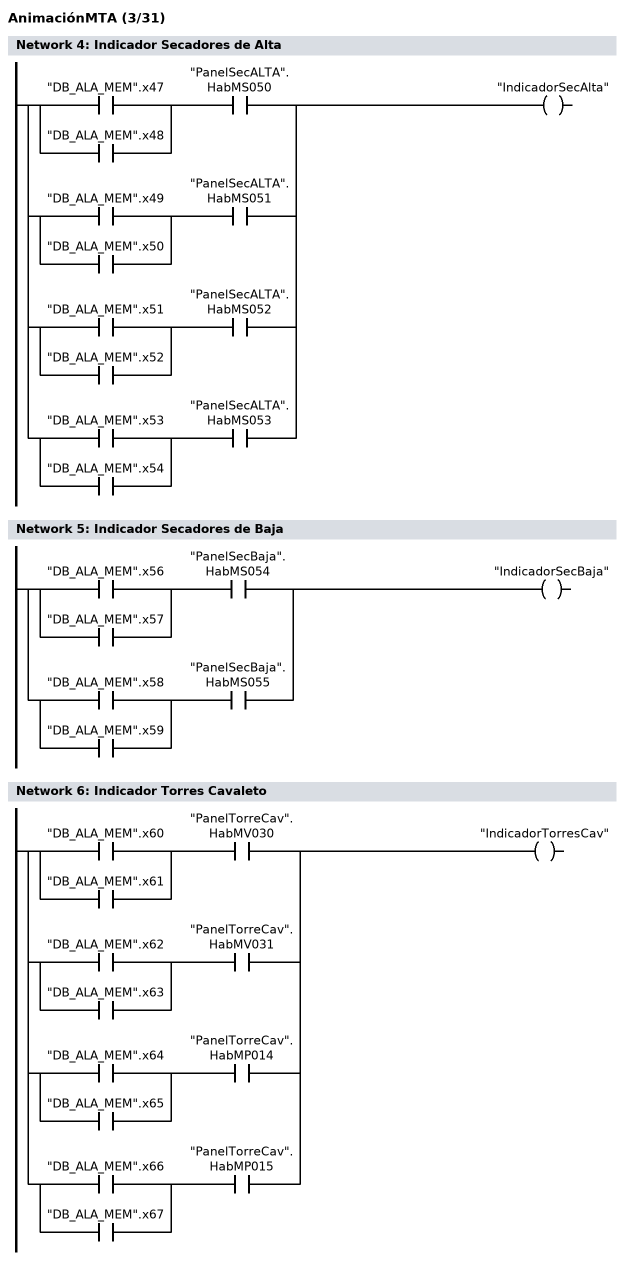
   RUNG wire#powerrail
      Contact( "DB_ALA_MEM".x47 )
      wire#w1
      Contact( "PanelSecALTA".HabMS050 )
      wire#w2
      Coil( "IndicadorSecAlta" )
   END_RUNG
   RUNG wire#powerrail
      Contact( "DB_ALA_MEM".x48 )
   END_RUNG wire#w1
   RUNG wire#powerrail
      Contact( "DB_ALA_MEM".x49 )
      wire#w3
      Contact( "PanelSecALTA".HabMS051 )
   END_RUNG wire#w2
   RUNG wire#powerrail
      Contact( "DB_ALA_MEM".x50 )
   END_RUNG wire#w3
   RUNG wire#powerrail
      Contact( "DB_ALA_MEM".x51 )
      wire#w4
      Contact( "PanelSecALTA".HabMS052 )
   END_RUNG wire#w2
   RUNG wire#powerrail
      Contact( "DB_ALA_MEM".x52 )
   END_RUNG wire#w4
   RUNG wire#powerrail
      Contact( "DB_ALA_MEM".x53 )
      wire#w5
      Contact( "PanelSecALTA".HabMS053 )
   END_RUNG wire#w2
   RUNG wire#powerrail
      Contact( "DB_ALA_MEM".x54 )
   END_RUNG wire#w5
   // the same network as SCL:
   "IndicadorSecAlta" := (("DB_ALA_MEM".x47 OR "DB_ALA_MEM".x48) AND "PanelSecALTA".HabMS050) OR (("DB_ALA_MEM".x49 OR "DB_ALA_MEM".x50) AND "PanelSecALTA".HabMS051) OR (("DB_ALA_MEM".x51 OR "DB_ALA_MEM".x52) AND "PanelSecALTA".HabMS052) OR (("DB_ALA_MEM".x53 OR "DB_ALA_MEM".x54) AND "PanelSecALTA".HabMS053);
END_REGION

REGION Network 5: Indicador Secadores de Baja
   RUNG wire#powerrail
      Contact( "DB_ALA_MEM".x56 )
      wire#w1
      Contact( "PanelSecBaja".HabMS054 )
      wire#w2
      Coil( "IndicadorSecBaja" )
   END_RUNG
   RUNG wire#powerrail
      Contact( "DB_ALA_MEM".x57 )
   END_RUNG wire#w1
   RUNG wire#powerrail
      Contact( "DB_ALA_MEM".x58 )
      wire#w3
      Contact( "PanelSecBaja".HabMS055 )
   END_RUNG wire#w2
   RUNG wire#powerrail
      Contact( "DB_ALA_MEM".x59 )
   END_RUNG wire#w3
   // the same network as SCL:
   "IndicadorSecBaja" := (("DB_ALA_MEM".x56 OR "DB_ALA_MEM".x57) AND "PanelSecBaja".HabMS054) OR (("DB_ALA_MEM".x58 OR "DB_ALA_MEM".x59) AND "PanelSecBaja".HabMS055);
END_REGION

REGION Network 6: Indicador Torres Cavaleto
   RUNG wire#powerrail
      Contact( "DB_ALA_MEM".x60 )
      wire#w1
      Contact( "PanelTorreCav".HabMV030 )
      wire#w2
      Coil( "IndicadorTorresCav" )
   END_RUNG
   RUNG wire#powerrail
      Contact( "DB_ALA_MEM".x61 )
   END_RUNG wire#w1
   RUNG wire#powerrail
      Contact( "DB_ALA_MEM".x62 )
      wire#w3
      Contact( "PanelTorreCav".HabMV031 )
   END_RUNG wire#w2
   RUNG wire#powerrail
      Contact( "DB_ALA_MEM".x63 )
   END_RUNG wire#w3
   RUNG wire#powerrail
      Contact( "DB_ALA_MEM".x64 )
      wire#w4
      Contact( "PanelTorreCav".HabMP014 )
   END_RUNG wire#w2
   RUNG wire#powerrail
      Contact( "DB_ALA_MEM".x65 )
   END_RUNG wire#w4
   RUNG wire#powerrail
      Contact( "DB_ALA_MEM".x66 )
      wire#w5
      Contact( "PanelTorreCav".HabMP015 )
   END_RUNG wire#w2
   RUNG wire#powerrail
      Contact( "DB_ALA_MEM".x67 )
   END_RUNG wire#w5
   // the same network as SCL:
   "IndicadorTorresCav" := (("DB_ALA_MEM".x60 OR "DB_ALA_MEM".x61) AND "PanelTorreCav".HabMV030) OR (("DB_ALA_MEM".x62 OR "DB_ALA_MEM".x63) AND "PanelTorreCav".HabMV031) OR (("DB_ALA_MEM".x64 OR "DB_ALA_MEM".x65) AND "PanelTorreCav".HabMP014) OR (("DB_ALA_MEM".x66 OR "DB_ALA_MEM".x67) AND "PanelTorreCav".HabMP015);
END_REGION

REGION Network 7: Indicador Compresores de Alta
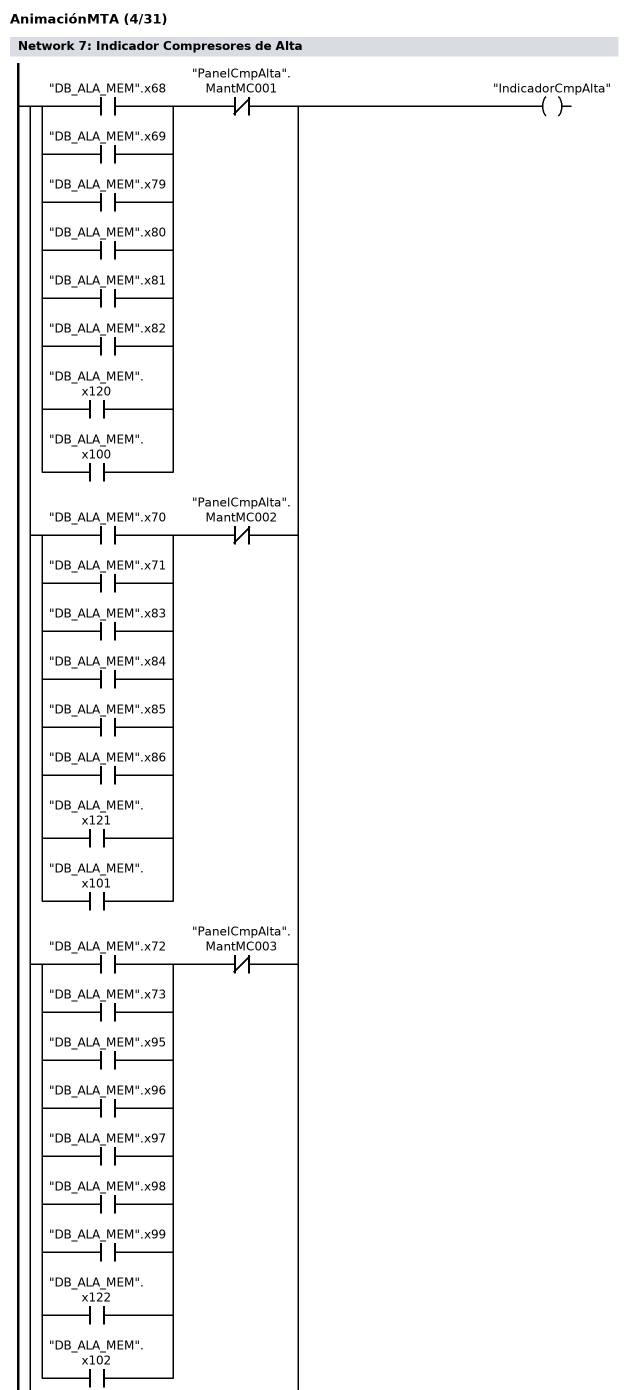
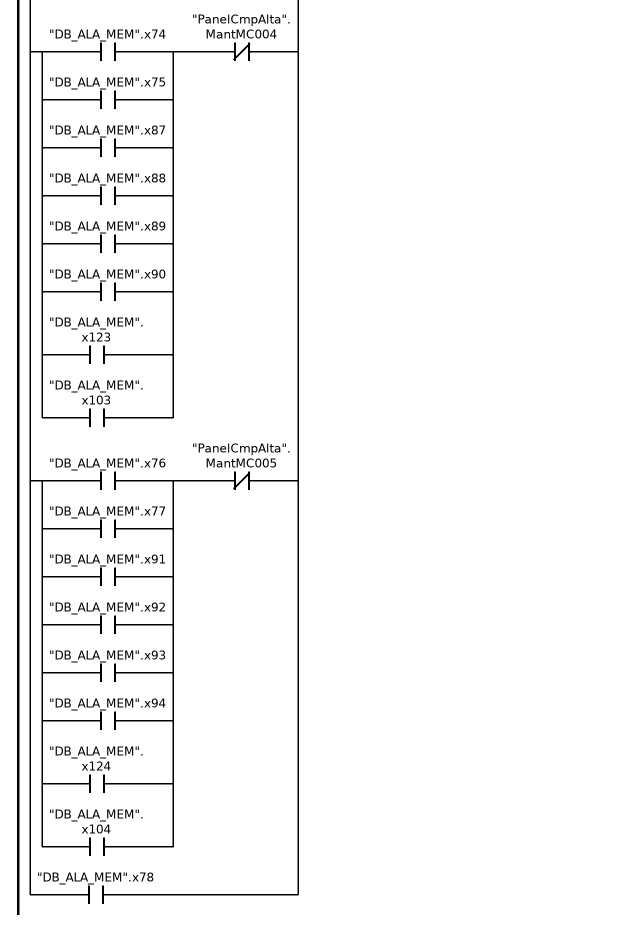
   RUNG wire#powerrail
      Contact( "DB_ALA_MEM".x68 )
      wire#w1
      I_Contact( "PanelCmpAlta".MantMC001 )
      wire#w2
      Coil( "IndicadorCmpAlta" )
   END_RUNG
   RUNG wire#powerrail
      Contact( "DB_ALA_MEM".x69 )
   END_RUNG wire#w1
   RUNG wire#powerrail
      Contact( "DB_ALA_MEM".x79 )
   END_RUNG wire#w1
   RUNG wire#powerrail
      Contact( "DB_ALA_MEM".x80 )
   END_RUNG wire#w1
   RUNG wire#powerrail
      Contact( "DB_ALA_MEM".x81 )
   END_RUNG wire#w1
   RUNG wire#powerrail
      Contact( "DB_ALA_MEM".x82 )
   END_RUNG wire#w1
   RUNG wire#powerrail
      Contact( "DB_ALA_MEM".x120 )
   END_RUNG wire#w1
   RUNG wire#powerrail
      Contact( "DB_ALA_MEM".x100 )
   END_RUNG wire#w1
   RUNG wire#powerrail
      Contact( "DB_ALA_MEM".x70 )
      wire#w3
      I_Contact( "PanelCmpAlta".MantMC002 )
   END_RUNG wire#w2
   RUNG wire#powerrail
      Contact( "DB_ALA_MEM".x71 )
   END_RUNG wire#w3
   RUNG wire#powerrail
      Contact( "DB_ALA_MEM".x83 )
   END_RUNG wire#w3
   RUNG wire#powerrail
      Contact( "DB_ALA_MEM".x84 )
   END_RUNG wire#w3
   RUNG wire#powerrail
      Contact( "DB_ALA_MEM".x85 )
   END_RUNG wire#w3
   RUNG wire#powerrail
      Contact( "DB_ALA_MEM".x86 )
   END_RUNG wire#w3
   RUNG wire#powerrail
      Contact( "DB_ALA_MEM".x121 )
   END_RUNG wire#w3
   RUNG wire#powerrail
      Contact( "DB_ALA_MEM".x101 )
   END_RUNG wire#w3
   RUNG wire#powerrail
      Contact( "DB_ALA_MEM".x72 )
      wire#w4
      I_Contact( "PanelCmpAlta".MantMC003 )
   END_RUNG wire#w2
   RUNG wire#powerrail
      Contact( "DB_ALA_MEM".x73 )
   END_RUNG wire#w4
   RUNG wire#powerrail
      Contact( "DB_ALA_MEM".x95 )
   END_RUNG wire#w4
   RUNG wire#powerrail
      Contact( "DB_ALA_MEM".x96 )
   END_RUNG wire#w4
   RUNG wire#powerrail
      Contact( "DB_ALA_MEM".x97 )
   END_RUNG wire#w4
   RUNG wire#powerrail
      Contact( "DB_ALA_MEM".x98 )
   END_RUNG wire#w4
   RUNG wire#powerrail
      Contact( "DB_ALA_MEM".x99 )
   END_RUNG wire#w4
   RUNG wire#powerrail
      Contact( "DB_ALA_MEM".x122 )
   END_RUNG wire#w4
   RUNG wire#powerrail
      Contact( "DB_ALA_MEM".x102 )
   END_RUNG wire#w4
   RUNG wire#powerrail
      Contact( "DB_ALA_MEM".x74 )
      wire#w5
      I_Contact( "PanelCmpAlta".MantMC004 )
   END_RUNG wire#w2
   RUNG wire#powerrail
      Contact( "DB_ALA_MEM".x75 )
   END_RUNG wire#w5
   RUNG wire#powerrail
      Contact( "DB_ALA_MEM".x87 )
   END_RUNG wire#w5
   RUNG wire#powerrail
      Contact( "DB_ALA_MEM".x88 )
   END_RUNG wire#w5
   RUNG wire#powerrail
      Contact( "DB_ALA_MEM".x89 )
   END_RUNG wire#w5
   RUNG wire#powerrail
      Contact( "DB_ALA_MEM".x90 )
   END_RUNG wire#w5
   RUNG wire#powerrail
      Contact( "DB_ALA_MEM".x123 )
   END_RUNG wire#w5
   RUNG wire#powerrail
      Contact( "DB_ALA_MEM".x103 )
   END_RUNG wire#w5
   RUNG wire#powerrail
      Contact( "DB_ALA_MEM".x76 )
      wire#w6
      I_Contact( "PanelCmpAlta".MantMC005 )
   END_RUNG wire#w2
   RUNG wire#powerrail
      Contact( "DB_ALA_MEM".x77 )
   END_RUNG wire#w6
   RUNG wire#powerrail
      Contact( "DB_ALA_MEM".x91 )
   END_RUNG wire#w6
   RUNG wire#powerrail
      Contact( "DB_ALA_MEM".x92 )
   END_RUNG wire#w6
   RUNG wire#powerrail
      Contact( "DB_ALA_MEM".x93 )
   END_RUNG wire#w6
   RUNG wire#powerrail
      Contact( "DB_ALA_MEM".x94 )
   END_RUNG wire#w6
   RUNG wire#powerrail
      Contact( "DB_ALA_MEM".x124 )
   END_RUNG wire#w6
   RUNG wire#powerrail
      Contact( "DB_ALA_MEM".x104 )
   END_RUNG wire#w6
   RUNG wire#powerrail
      Contact( "DB_ALA_MEM".x78 )
   END_RUNG wire#w2
   // the same network as SCL:
   "IndicadorCmpAlta" := (("DB_ALA_MEM".x68 OR "DB_ALA_MEM".x69 OR "DB_ALA_MEM".x79 OR "DB_ALA_MEM".x80 OR "DB_ALA_MEM".x81 OR "DB_ALA_MEM".x82 OR "DB_ALA_MEM".x120 OR "DB_ALA_MEM".x100) AND NOT "PanelCmpAlta".MantMC001) OR (("DB_ALA_MEM".x70 OR "DB_ALA_MEM".x71 OR "DB_ALA_MEM".x83 OR "DB_ALA_MEM".x84 OR "DB_ALA_MEM".x85 OR "DB_ALA_MEM".x86 OR "DB_ALA_MEM".x121 OR "DB_ALA_MEM".x101) AND NOT "PanelCmpAlta".MantMC002) OR (("DB_ALA_MEM".x72 OR "DB_ALA_MEM".x73 OR "DB_ALA_MEM".x95 OR "DB_ALA_MEM".x96 OR "DB_ALA_MEM".x97 OR "DB_ALA_MEM".x98 OR "DB_ALA_MEM".x99 OR "DB_ALA_MEM".x122 OR "DB_ALA_MEM".x102) AND NOT "PanelCmpAlta".MantMC003) OR (("DB_ALA_MEM".x74 OR "DB_ALA_MEM".x75 OR "DB_ALA_MEM".x87 OR "DB_ALA_MEM".x88 OR "DB_ALA_MEM".x89 OR "DB_ALA_MEM".x90 OR "DB_ALA_MEM".x123 OR "DB_ALA_MEM".x103) AND NOT "PanelCmpAlta".MantMC004) OR (("DB_ALA_MEM".x76 OR "DB_ALA_MEM".x77 OR "DB_ALA_MEM".x91 OR "DB_ALA_MEM".x92 OR "DB_ALA_MEM".x93 OR "DB_ALA_MEM".x94 OR "DB_ALA_MEM".x124 OR "DB_ALA_MEM".x104) AND NOT "PanelCmpAlta".MantMC005) OR "DB_ALA_MEM".x78;
END_REGION

REGION Network 8: Animación MT007 - Bomba Intercambiador LÍNEA 1
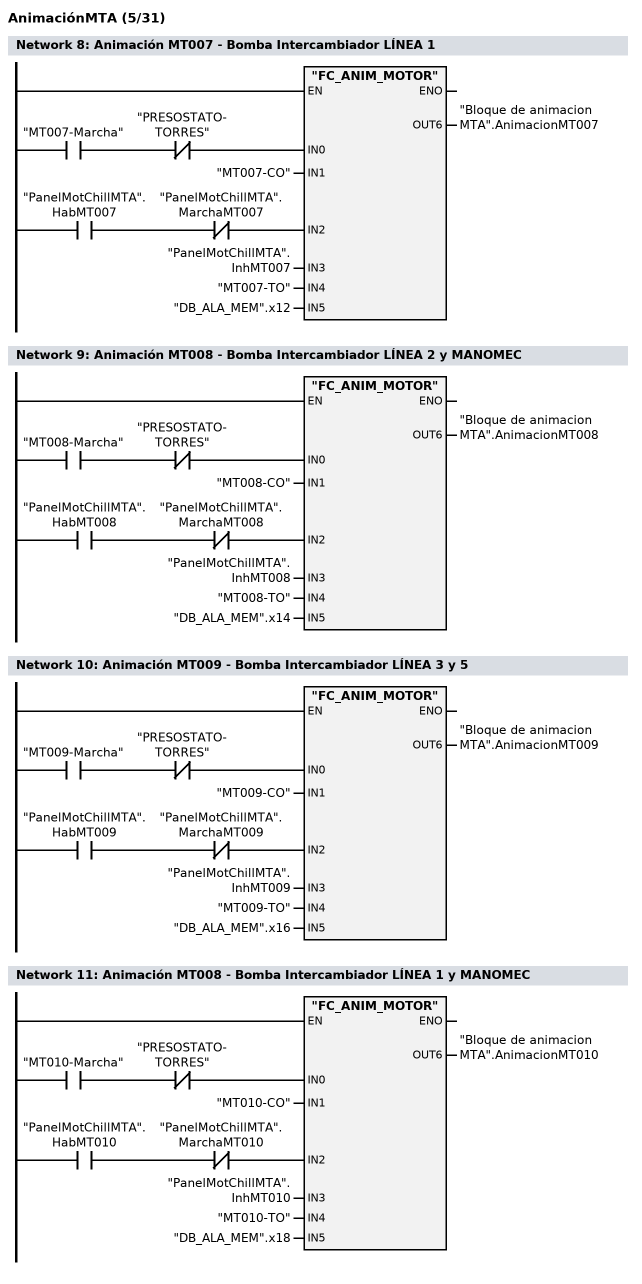
   RUNG wire#powerrail
      "FC_ANIM_MOTOR"(IN0 := wire#w1, IN2 := wire#w2, IN1 := "MT007-CO", IN3 := "PanelMotChillMTA".InhMT007, IN4 := "MT007-TO", IN5 := "DB_ALA_MEM".x12, OUT6 => "Bloque de animacion MTA".AnimacionMT007)
   END_RUNG
   RUNG wire#powerrail
      Contact( "MT007-Marcha" )
      I_Contact( "PRESOSTATO-TORRES" )
   END_RUNG wire#w1
   RUNG wire#powerrail
      Contact( "PanelMotChillMTA".HabMT007 )
      I_Contact( "PanelMotChillMTA".MarchaMT007 )
   END_RUNG wire#w2
   // the same network as SCL:
   "FC_ANIM_MOTOR"(IN0 := "MT007-Marcha" AND NOT "PRESOSTATO-TORRES",
                   IN1 := "MT007-CO",
                   IN2 := "PanelMotChillMTA".HabMT007 AND NOT "PanelMotChillMTA".MarchaMT007,
                   IN3 := "PanelMotChillMTA".InhMT007,
                   IN4 := "MT007-TO",
                   IN5 := "DB_ALA_MEM".x12,
                   OUT6 => "Bloque de animacion MTA".AnimacionMT007);
END_REGION

REGION Network 9: Animación MT008 - Bomba Intercambiador LÍNEA 2 y MANOMEC
   RUNG wire#powerrail
      "FC_ANIM_MOTOR"(IN0 := wire#w1, IN2 := wire#w2, IN1 := "MT008-CO", IN3 := "PanelMotChillMTA".InhMT008, IN4 := "MT008-TO", IN5 := "DB_ALA_MEM".x14, OUT6 => "Bloque de animacion MTA".AnimacionMT008)
   END_RUNG
   RUNG wire#powerrail
      Contact( "MT008-Marcha" )
      I_Contact( "PRESOSTATO-TORRES" )
   END_RUNG wire#w1
   RUNG wire#powerrail
      Contact( "PanelMotChillMTA".HabMT008 )
      I_Contact( "PanelMotChillMTA".MarchaMT008 )
   END_RUNG wire#w2
   // the same network as SCL:
   "FC_ANIM_MOTOR"(IN0 := "MT008-Marcha" AND NOT "PRESOSTATO-TORRES",
                   IN1 := "MT008-CO",
                   IN2 := "PanelMotChillMTA".HabMT008 AND NOT "PanelMotChillMTA".MarchaMT008,
                   IN3 := "PanelMotChillMTA".InhMT008,
                   IN4 := "MT008-TO",
                   IN5 := "DB_ALA_MEM".x14,
                   OUT6 => "Bloque de animacion MTA".AnimacionMT008);
END_REGION

REGION Network 10: Animación MT009 - Bomba Intercambiador LÍNEA 3 y 5
   RUNG wire#powerrail
      "FC_ANIM_MOTOR"(IN0 := wire#w1, IN2 := wire#w2, IN1 := "MT009-CO", IN3 := "PanelMotChillMTA".InhMT009, IN4 := "MT009-TO", IN5 := "DB_ALA_MEM".x16, OUT6 => "Bloque de animacion MTA".AnimacionMT009)
   END_RUNG
   RUNG wire#powerrail
      Contact( "MT009-Marcha" )
      I_Contact( "PRESOSTATO-TORRES" )
   END_RUNG wire#w1
   RUNG wire#powerrail
      Contact( "PanelMotChillMTA".HabMT009 )
      I_Contact( "PanelMotChillMTA".MarchaMT009 )
   END_RUNG wire#w2
   // the same network as SCL:
   "FC_ANIM_MOTOR"(IN0 := "MT009-Marcha" AND NOT "PRESOSTATO-TORRES",
                   IN1 := "MT009-CO",
                   IN2 := "PanelMotChillMTA".HabMT009 AND NOT "PanelMotChillMTA".MarchaMT009,
                   IN3 := "PanelMotChillMTA".InhMT009,
                   IN4 := "MT009-TO",
                   IN5 := "DB_ALA_MEM".x16,
                   OUT6 => "Bloque de animacion MTA".AnimacionMT009);
END_REGION

REGION Network 11: Animación MT008 - Bomba Intercambiador LÍNEA 1 y MANOMEC
   RUNG wire#powerrail
      "FC_ANIM_MOTOR"(IN0 := wire#w1, IN2 := wire#w2, IN1 := "MT010-CO", IN3 := "PanelMotChillMTA".InhMT010, IN4 := "MT010-TO", IN5 := "DB_ALA_MEM".x18, OUT6 => "Bloque de animacion MTA".AnimacionMT010)
   END_RUNG
   RUNG wire#powerrail
      Contact( "MT010-Marcha" )
      I_Contact( "PRESOSTATO-TORRES" )
   END_RUNG wire#w1
   RUNG wire#powerrail
      Contact( "PanelMotChillMTA".HabMT010 )
      I_Contact( "PanelMotChillMTA".MarchaMT010 )
   END_RUNG wire#w2
   // the same network as SCL:
   "FC_ANIM_MOTOR"(IN0 := "MT010-Marcha" AND NOT "PRESOSTATO-TORRES",
                   IN1 := "MT010-CO",
                   IN2 := "PanelMotChillMTA".HabMT010 AND NOT "PanelMotChillMTA".MarchaMT010,
                   IN3 := "PanelMotChillMTA".InhMT010,
                   IN4 := "MT010-TO",
                   IN5 := "DB_ALA_MEM".x18,
                   OUT6 => "Bloque de animacion MTA".AnimacionMT010);
END_REGION

REGION Network 12: Animación MP010 - Bomba Principal Chillers Soplado
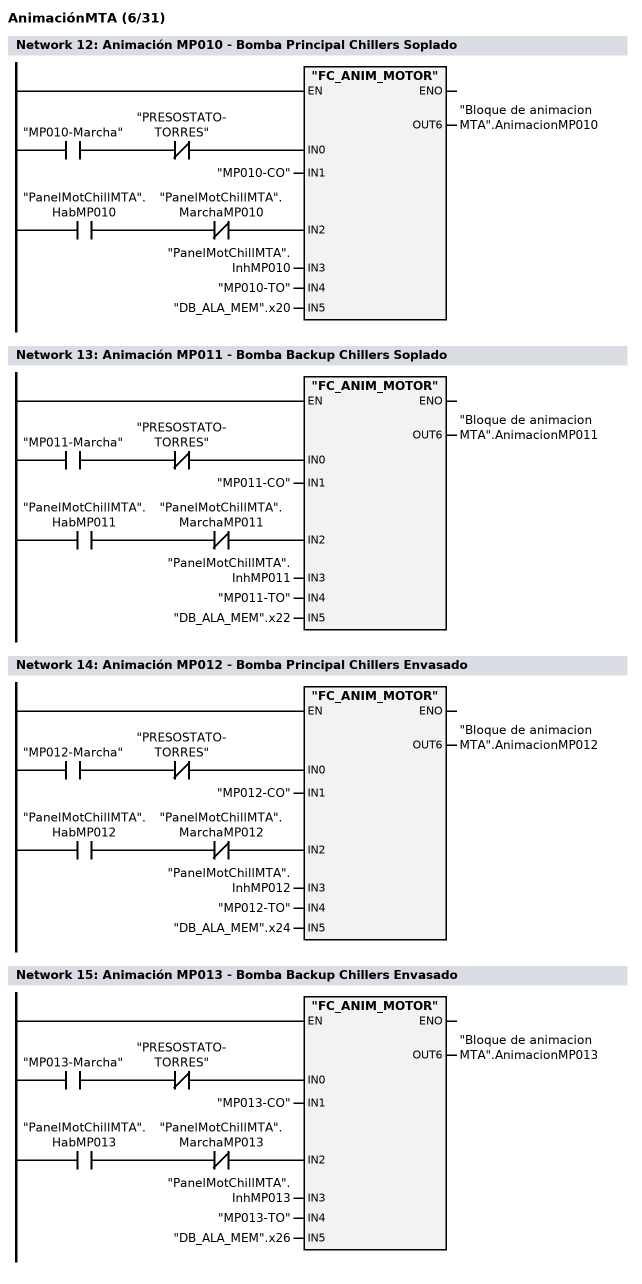
   RUNG wire#powerrail
      "FC_ANIM_MOTOR"(IN0 := wire#w1, IN2 := wire#w2, IN1 := "MP010-CO", IN3 := "PanelMotChillMTA".InhMP010, IN4 := "MP010-TO", IN5 := "DB_ALA_MEM".x20, OUT6 => "Bloque de animacion MTA".AnimacionMP010)
   END_RUNG
   RUNG wire#powerrail
      Contact( "MP010-Marcha" )
      I_Contact( "PRESOSTATO-TORRES" )
   END_RUNG wire#w1
   RUNG wire#powerrail
      Contact( "PanelMotChillMTA".HabMP010 )
      I_Contact( "PanelMotChillMTA".MarchaMP010 )
   END_RUNG wire#w2
   // the same network as SCL:
   "FC_ANIM_MOTOR"(IN0 := "MP010-Marcha" AND NOT "PRESOSTATO-TORRES",
                   IN1 := "MP010-CO",
                   IN2 := "PanelMotChillMTA".HabMP010 AND NOT "PanelMotChillMTA".MarchaMP010,
                   IN3 := "PanelMotChillMTA".InhMP010,
                   IN4 := "MP010-TO",
                   IN5 := "DB_ALA_MEM".x20,
                   OUT6 => "Bloque de animacion MTA".AnimacionMP010);
END_REGION

REGION Network 13: Animación MP011 - Bomba Backup Chillers Soplado
   RUNG wire#powerrail
      "FC_ANIM_MOTOR"(IN0 := wire#w1, IN2 := wire#w2, IN1 := "MP011-CO", IN3 := "PanelMotChillMTA".InhMP011, IN4 := "MP011-TO", IN5 := "DB_ALA_MEM".x22, OUT6 => "Bloque de animacion MTA".AnimacionMP011)
   END_RUNG
   RUNG wire#powerrail
      Contact( "MP011-Marcha" )
      I_Contact( "PRESOSTATO-TORRES" )
   END_RUNG wire#w1
   RUNG wire#powerrail
      Contact( "PanelMotChillMTA".HabMP011 )
      I_Contact( "PanelMotChillMTA".MarchaMP011 )
   END_RUNG wire#w2
   // the same network as SCL:
   "FC_ANIM_MOTOR"(IN0 := "MP011-Marcha" AND NOT "PRESOSTATO-TORRES",
                   IN1 := "MP011-CO",
                   IN2 := "PanelMotChillMTA".HabMP011 AND NOT "PanelMotChillMTA".MarchaMP011,
                   IN3 := "PanelMotChillMTA".InhMP011,
                   IN4 := "MP011-TO",
                   IN5 := "DB_ALA_MEM".x22,
                   OUT6 => "Bloque de animacion MTA".AnimacionMP011);
END_REGION

REGION Network 14: Animación MP012 - Bomba Principal Chillers Envasado
   RUNG wire#powerrail
      "FC_ANIM_MOTOR"(IN0 := wire#w1, IN2 := wire#w2, IN1 := "MP012-CO", IN3 := "PanelMotChillMTA".InhMP012, IN4 := "MP012-TO", IN5 := "DB_ALA_MEM".x24, OUT6 => "Bloque de animacion MTA".AnimacionMP012)
   END_RUNG
   RUNG wire#powerrail
      Contact( "MP012-Marcha" )
      I_Contact( "PRESOSTATO-TORRES" )
   END_RUNG wire#w1
   RUNG wire#powerrail
      Contact( "PanelMotChillMTA".HabMP012 )
      I_Contact( "PanelMotChillMTA".MarchaMP012 )
   END_RUNG wire#w2
   // the same network as SCL:
   "FC_ANIM_MOTOR"(IN0 := "MP012-Marcha" AND NOT "PRESOSTATO-TORRES",
                   IN1 := "MP012-CO",
                   IN2 := "PanelMotChillMTA".HabMP012 AND NOT "PanelMotChillMTA".MarchaMP012,
                   IN3 := "PanelMotChillMTA".InhMP012,
                   IN4 := "MP012-TO",
                   IN5 := "DB_ALA_MEM".x24,
                   OUT6 => "Bloque de animacion MTA".AnimacionMP012);
END_REGION

REGION Network 15: Animación MP013 - Bomba Backup Chillers Envasado
   RUNG wire#powerrail
      "FC_ANIM_MOTOR"(IN0 := wire#w1, IN2 := wire#w2, IN1 := "MP013-CO", IN3 := "PanelMotChillMTA".InhMP013, IN4 := "MP013-TO", IN5 := "DB_ALA_MEM".x26, OUT6 => "Bloque de animacion MTA".AnimacionMP013)
   END_RUNG
   RUNG wire#powerrail
      Contact( "MP013-Marcha" )
      I_Contact( "PRESOSTATO-TORRES" )
   END_RUNG wire#w1
   RUNG wire#powerrail
      Contact( "PanelMotChillMTA".HabMP013 )
      I_Contact( "PanelMotChillMTA".MarchaMP013 )
   END_RUNG wire#w2
   // the same network as SCL:
   "FC_ANIM_MOTOR"(IN0 := "MP013-Marcha" AND NOT "PRESOSTATO-TORRES",
                   IN1 := "MP013-CO",
                   IN2 := "PanelMotChillMTA".HabMP013 AND NOT "PanelMotChillMTA".MarchaMP013,
                   IN3 := "PanelMotChillMTA".InhMP013,
                   IN4 := "MP013-TO",
                   IN5 := "DB_ALA_MEM".x26,
                   OUT6 => "Bloque de animacion MTA".AnimacionMP013);
END_REGION

REGION Network 16: Animación MP018 - Bomba 1 Torres de enfriamiento
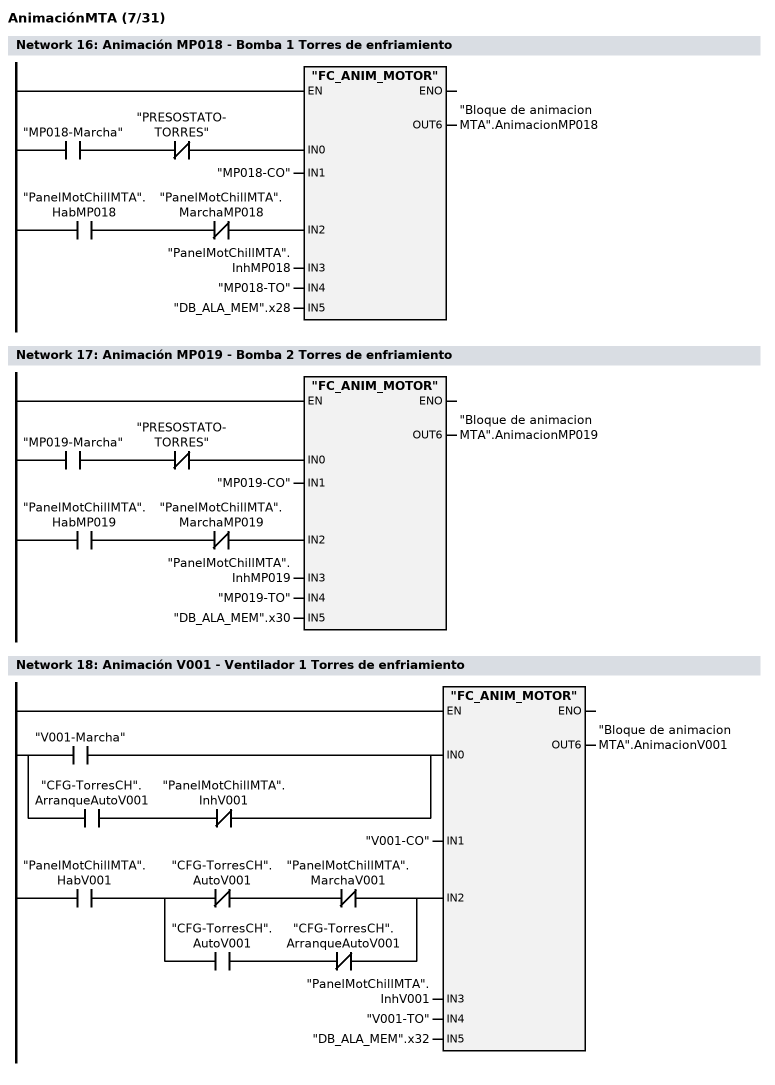
   RUNG wire#powerrail
      "FC_ANIM_MOTOR"(IN0 := wire#w1, IN2 := wire#w2, IN1 := "MP018-CO", IN3 := "PanelMotChillMTA".InhMP018, IN4 := "MP018-TO", IN5 := "DB_ALA_MEM".x28, OUT6 => "Bloque de animacion MTA".AnimacionMP018)
   END_RUNG
   RUNG wire#powerrail
      Contact( "MP018-Marcha" )
      I_Contact( "PRESOSTATO-TORRES" )
   END_RUNG wire#w1
   RUNG wire#powerrail
      Contact( "PanelMotChillMTA".HabMP018 )
      I_Contact( "PanelMotChillMTA".MarchaMP018 )
   END_RUNG wire#w2
   // the same network as SCL:
   "FC_ANIM_MOTOR"(IN0 := "MP018-Marcha" AND NOT "PRESOSTATO-TORRES",
                   IN1 := "MP018-CO",
                   IN2 := "PanelMotChillMTA".HabMP018 AND NOT "PanelMotChillMTA".MarchaMP018,
                   IN3 := "PanelMotChillMTA".InhMP018,
                   IN4 := "MP018-TO",
                   IN5 := "DB_ALA_MEM".x28,
                   OUT6 => "Bloque de animacion MTA".AnimacionMP018);
END_REGION

REGION Network 17: Animación MP019 - Bomba 2 Torres de enfriamiento
   RUNG wire#powerrail
      "FC_ANIM_MOTOR"(IN0 := wire#w1, IN2 := wire#w2, IN1 := "MP019-CO", IN3 := "PanelMotChillMTA".InhMP019, IN4 := "MP019-TO", IN5 := "DB_ALA_MEM".x30, OUT6 => "Bloque de animacion MTA".AnimacionMP019)
   END_RUNG
   RUNG wire#powerrail
      Contact( "MP019-Marcha" )
      I_Contact( "PRESOSTATO-TORRES" )
   END_RUNG wire#w1
   RUNG wire#powerrail
      Contact( "PanelMotChillMTA".HabMP019 )
      I_Contact( "PanelMotChillMTA".MarchaMP019 )
   END_RUNG wire#w2
   // the same network as SCL:
   "FC_ANIM_MOTOR"(IN0 := "MP019-Marcha" AND NOT "PRESOSTATO-TORRES",
                   IN1 := "MP019-CO",
                   IN2 := "PanelMotChillMTA".HabMP019 AND NOT "PanelMotChillMTA".MarchaMP019,
                   IN3 := "PanelMotChillMTA".InhMP019,
                   IN4 := "MP019-TO",
                   IN5 := "DB_ALA_MEM".x30,
                   OUT6 => "Bloque de animacion MTA".AnimacionMP019);
END_REGION

REGION Network 18: Animación V001 - Ventilador 1 Torres de enfriamiento
   RUNG wire#powerrail
      "FC_ANIM_MOTOR"(IN0 := wire#w1, IN2 := wire#w3, IN1 := "V001-CO", IN3 := "PanelMotChillMTA".InhV001, IN4 := "V001-TO", IN5 := "DB_ALA_MEM".x32, OUT6 => "Bloque de animacion MTA".AnimacionV001)
   END_RUNG
   RUNG wire#powerrail
      Contact( "V001-Marcha" )
   END_RUNG wire#w1
   RUNG wire#powerrail
      Contact( "CFG-TorresCH".ArranqueAutoV001 )
      I_Contact( "PanelMotChillMTA".InhV001 )
   END_RUNG wire#w1
   RUNG wire#powerrail
      Contact( "PanelMotChillMTA".HabV001 )
      wire#w2
      I_Contact( "CFG-TorresCH".AutoV001 )
      I_Contact( "PanelMotChillMTA".MarchaV001 )
   END_RUNG wire#w3
   RUNG wire#w2
      Contact( "CFG-TorresCH".AutoV001 )
      I_Contact( "CFG-TorresCH".ArranqueAutoV001 )
   END_RUNG wire#w3
   // the same network as SCL:
   "FC_ANIM_MOTOR"(IN0 := "V001-Marcha" OR ("CFG-TorresCH".ArranqueAutoV001 AND NOT "PanelMotChillMTA".InhV001),
                   IN1 := "V001-CO",
                   IN2 := "PanelMotChillMTA".HabV001 AND ((NOT "CFG-TorresCH".AutoV001 AND NOT "PanelMotChillMTA".MarchaV001) OR ("CFG-TorresCH".AutoV001 AND NOT "CFG-TorresCH".ArranqueAutoV001)),
                   IN3 := "PanelMotChillMTA".InhV001,
                   IN4 := "V001-TO",
                   IN5 := "DB_ALA_MEM".x32,
                   OUT6 => "Bloque de animacion MTA".AnimacionV001);
END_REGION

REGION Network 19: Animación V002 - Ventilador 2 Torres de enfriamiento
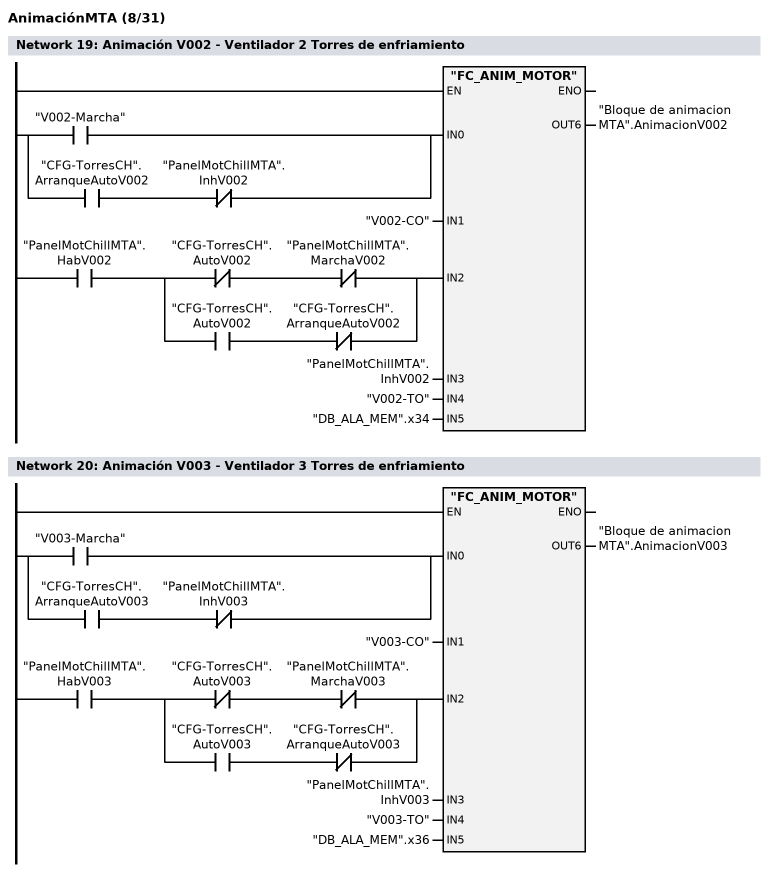
   RUNG wire#powerrail
      "FC_ANIM_MOTOR"(IN0 := wire#w1, IN2 := wire#w3, IN1 := "V002-CO", IN3 := "PanelMotChillMTA".InhV002, IN4 := "V002-TO", IN5 := "DB_ALA_MEM".x34, OUT6 => "Bloque de animacion MTA".AnimacionV002)
   END_RUNG
   RUNG wire#powerrail
      Contact( "V002-Marcha" )
   END_RUNG wire#w1
   RUNG wire#powerrail
      Contact( "CFG-TorresCH".ArranqueAutoV002 )
      I_Contact( "PanelMotChillMTA".InhV002 )
   END_RUNG wire#w1
   RUNG wire#powerrail
      Contact( "PanelMotChillMTA".HabV002 )
      wire#w2
      I_Contact( "CFG-TorresCH".AutoV002 )
      I_Contact( "PanelMotChillMTA".MarchaV002 )
   END_RUNG wire#w3
   RUNG wire#w2
      Contact( "CFG-TorresCH".AutoV002 )
      I_Contact( "CFG-TorresCH".ArranqueAutoV002 )
   END_RUNG wire#w3
   // the same network as SCL:
   "FC_ANIM_MOTOR"(IN0 := "V002-Marcha" OR ("CFG-TorresCH".ArranqueAutoV002 AND NOT "PanelMotChillMTA".InhV002),
                   IN1 := "V002-CO",
                   IN2 := "PanelMotChillMTA".HabV002 AND ((NOT "CFG-TorresCH".AutoV002 AND NOT "PanelMotChillMTA".MarchaV002) OR ("CFG-TorresCH".AutoV002 AND NOT "CFG-TorresCH".ArranqueAutoV002)),
                   IN3 := "PanelMotChillMTA".InhV002,
                   IN4 := "V002-TO",
                   IN5 := "DB_ALA_MEM".x34,
                   OUT6 => "Bloque de animacion MTA".AnimacionV002);
END_REGION

REGION Network 20: Animación V003 - Ventilador 3 Torres de enfriamiento
   RUNG wire#powerrail
      "FC_ANIM_MOTOR"(IN0 := wire#w1, IN2 := wire#w3, IN1 := "V003-CO", IN3 := "PanelMotChillMTA".InhV003, IN4 := "V003-TO", IN5 := "DB_ALA_MEM".x36, OUT6 => "Bloque de animacion MTA".AnimacionV003)
   END_RUNG
   RUNG wire#powerrail
      Contact( "V003-Marcha" )
   END_RUNG wire#w1
   RUNG wire#powerrail
      Contact( "CFG-TorresCH".ArranqueAutoV003 )
      I_Contact( "PanelMotChillMTA".InhV003 )
   END_RUNG wire#w1
   RUNG wire#powerrail
      Contact( "PanelMotChillMTA".HabV003 )
      wire#w2
      I_Contact( "CFG-TorresCH".AutoV003 )
      I_Contact( "PanelMotChillMTA".MarchaV003 )
   END_RUNG wire#w3
   RUNG wire#w2
      Contact( "CFG-TorresCH".AutoV003 )
      I_Contact( "CFG-TorresCH".ArranqueAutoV003 )
   END_RUNG wire#w3
   // the same network as SCL:
   "FC_ANIM_MOTOR"(IN0 := "V003-Marcha" OR ("CFG-TorresCH".ArranqueAutoV003 AND NOT "PanelMotChillMTA".InhV003),
                   IN1 := "V003-CO",
                   IN2 := "PanelMotChillMTA".HabV003 AND ((NOT "CFG-TorresCH".AutoV003 AND NOT "PanelMotChillMTA".MarchaV003) OR ("CFG-TorresCH".AutoV003 AND NOT "CFG-TorresCH".ArranqueAutoV003)),
                   IN3 := "PanelMotChillMTA".InhV003,
                   IN4 := "V003-TO",
                   IN5 := "DB_ALA_MEM".x36,
                   OUT6 => "Bloque de animacion MTA".AnimacionV003);
END_REGION

REGION Network 21: Animación MC060 - Compresor de Baja SULLAIR 2
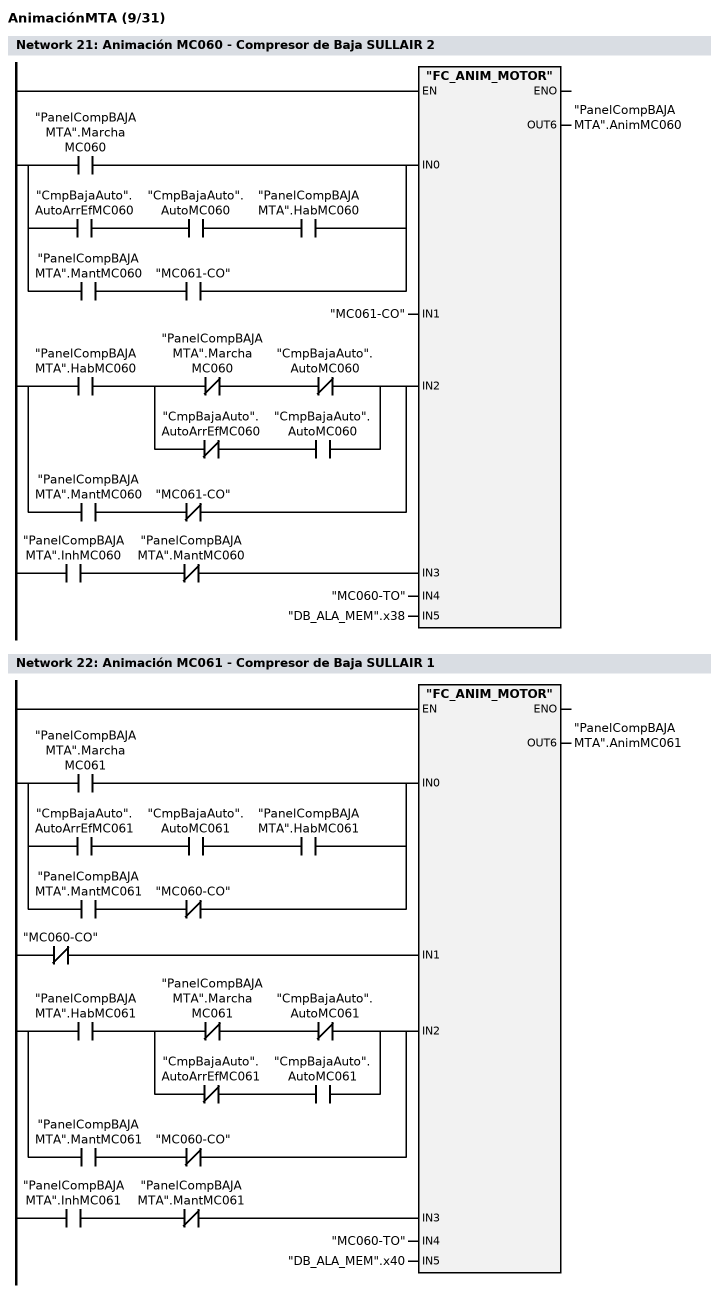
   RUNG wire#powerrail
      "FC_ANIM_MOTOR"(IN0 := wire#w1, IN2 := wire#w3, IN3 := wire#w4, IN1 := "MC061-CO", IN4 := "MC060-TO", IN5 := "DB_ALA_MEM".x38, OUT6 => "PanelCompBAJA MTA".AnimMC060)
   END_RUNG
   RUNG wire#powerrail
      Contact( "PanelCompBAJA MTA".MarchaMC060 )
   END_RUNG wire#w1
   RUNG wire#powerrail
      Contact( "CmpBajaAuto".AutoArrEfMC060 )
      Contact( "CmpBajaAuto".AutoMC060 )
      Contact( "PanelCompBAJA MTA".HabMC060 )
   END_RUNG wire#w1
   RUNG wire#powerrail
      Contact( "PanelCompBAJA MTA".MantMC060 )
      Contact( "MC061-CO" )
   END_RUNG wire#w1
   RUNG wire#powerrail
      Contact( "PanelCompBAJA MTA".HabMC060 )
      wire#w2
      I_Contact( "PanelCompBAJA MTA".MarchaMC060 )
      I_Contact( "CmpBajaAuto".AutoMC060 )
   END_RUNG wire#w3
   RUNG wire#w2
      I_Contact( "CmpBajaAuto".AutoArrEfMC060 )
      Contact( "CmpBajaAuto".AutoMC060 )
   END_RUNG wire#w3
   RUNG wire#powerrail
      Contact( "PanelCompBAJA MTA".MantMC060 )
      I_Contact( "MC061-CO" )
   END_RUNG wire#w3
   RUNG wire#powerrail
      Contact( "PanelCompBAJA MTA".InhMC060 )
      I_Contact( "PanelCompBAJA MTA".MantMC060 )
   END_RUNG wire#w4
   // the same network as SCL:
   "FC_ANIM_MOTOR"(IN0 := "PanelCompBAJA MTA".MarchaMC060 OR ("CmpBajaAuto".AutoArrEfMC060 AND "CmpBajaAuto".AutoMC060 AND "PanelCompBAJA MTA".HabMC060) OR ("PanelCompBAJA MTA".MantMC060 AND "MC061-CO"),
                   IN1 := "MC061-CO",
                   IN2 := ("PanelCompBAJA MTA".HabMC060 AND ((NOT "PanelCompBAJA MTA".MarchaMC060 AND NOT "CmpBajaAuto".AutoMC060) OR (NOT "CmpBajaAuto".AutoArrEfMC060 AND "CmpBajaAuto".AutoMC060))) OR ("PanelCompBAJA MTA".MantMC060 AND NOT "MC061-CO"),
                   IN3 := "PanelCompBAJA MTA".InhMC060 AND NOT "PanelCompBAJA MTA".MantMC060,
                   IN4 := "MC060-TO",
                   IN5 := "DB_ALA_MEM".x38,
                   OUT6 => "PanelCompBAJA MTA".AnimMC060);
END_REGION

REGION Network 22: Animación MC061 - Compresor de Baja SULLAIR 1
   RUNG wire#powerrail
      "FC_ANIM_MOTOR"(IN0 := wire#w1, IN1 := wire#w2, IN2 := wire#w4, IN3 := wire#w5, IN4 := "MC060-TO", IN5 := "DB_ALA_MEM".x40, OUT6 => "PanelCompBAJA MTA".AnimMC061)
   END_RUNG
   RUNG wire#powerrail
      Contact( "PanelCompBAJA MTA".MarchaMC061 )
   END_RUNG wire#w1
   RUNG wire#powerrail
      Contact( "CmpBajaAuto".AutoArrEfMC061 )
      Contact( "CmpBajaAuto".AutoMC061 )
      Contact( "PanelCompBAJA MTA".HabMC061 )
   END_RUNG wire#w1
   RUNG wire#powerrail
      Contact( "PanelCompBAJA MTA".MantMC061 )
      I_Contact( "MC060-CO" )
   END_RUNG wire#w1
   RUNG wire#powerrail
      I_Contact( "MC060-CO" )
   END_RUNG wire#w2
   RUNG wire#powerrail
      Contact( "PanelCompBAJA MTA".HabMC061 )
      wire#w3
      I_Contact( "PanelCompBAJA MTA".MarchaMC061 )
      I_Contact( "CmpBajaAuto".AutoMC061 )
   END_RUNG wire#w4
   RUNG wire#w3
      I_Contact( "CmpBajaAuto".AutoArrEfMC061 )
      Contact( "CmpBajaAuto".AutoMC061 )
   END_RUNG wire#w4
   RUNG wire#powerrail
      Contact( "PanelCompBAJA MTA".MantMC061 )
      I_Contact( "MC060-CO" )
   END_RUNG wire#w4
   RUNG wire#powerrail
      Contact( "PanelCompBAJA MTA".InhMC061 )
      I_Contact( "PanelCompBAJA MTA".MantMC061 )
   END_RUNG wire#w5
   // the same network as SCL:
   "FC_ANIM_MOTOR"(IN0 := "PanelCompBAJA MTA".MarchaMC061 OR ("CmpBajaAuto".AutoArrEfMC061 AND "CmpBajaAuto".AutoMC061 AND "PanelCompBAJA MTA".HabMC061) OR ("PanelCompBAJA MTA".MantMC061 AND NOT "MC060-CO"),
                   IN1 := NOT "MC060-CO",
                   IN2 := ("PanelCompBAJA MTA".HabMC061 AND ((NOT "PanelCompBAJA MTA".MarchaMC061 AND NOT "CmpBajaAuto".AutoMC061) OR (NOT "CmpBajaAuto".AutoArrEfMC061 AND "CmpBajaAuto".AutoMC061))) OR ("PanelCompBAJA MTA".MantMC061 AND NOT "MC060-CO"),
                   IN3 := "PanelCompBAJA MTA".InhMC061 AND NOT "PanelCompBAJA MTA".MantMC061,
                   IN4 := "MC060-TO",
                   IN5 := "DB_ALA_MEM".x40,
                   OUT6 => "PanelCompBAJA MTA".AnimMC061);
END_REGION

REGION Network 23: Animación MC062 - Compresor de Baja SULLAIR 0
